                   REGION "INCREMENT FIRST STATION"
                       #firstStn += "simKP8Count";
                   END_REGION

                   REGION "UPPER LIMIT ROLL OVER"
                       IF #firstStn > "STATION_COUNT" THEN
                           #firstStn -= "STATION_COUNT" + 1;
                       END_IF;
                   END_REGION

               END_IF;
           END_REGION

           REGION "NEXT GROUP CHANGE DETECTION"
               #old.nextGrp := #currentBtn;
           END_REGION

       END_REGION

       REGION "PROCESS PREVIOUS GROUP PRESS"

           REGION "COPY TO LOCAL"
               #currentBtn := #simStations.up.actuate;
               #oldBtn := #old.prevGrp;
           END_REGION

           REGION "FALLING EDGE OF PREVIOUS GROUP"
               IF NOT #currentBtn AND #oldBtn THEN

                   REGION "DECREMENT FIRST STATION"
                       #firstStn -= "simKP8Count";
                   END_REGION

                   REGION "LOWER LIMIT ROLL OVER"
                       IF #firstStn < 0 THEN
                           #firstStn += "STATION_COUNT" + 1;
                       END_IF;
                   END_REGION

               END_IF;
           END_REGION

           REGION "PREVIOUS GROUP CHANGE DETECTION"
               #old.prevGrp := #currentBtn;
           END_REGION

       END_REGION

   END_REGION

   REGION "FOR EACH BUTTON"
       FOR #i := 0 TO 11 DO

           REGION "CALCULATE POINTER"
               #pStn := #i + #firstStn;
               #pSim := #i;
           END_REGION

           REGION "UPPER LIMIT ROLL OVER"
               IF #pStn > "STATION_COUNT" THEN
                   #pStn := #firstStn + #i - "STATION_COUNT" - 1;
               END_IF;
           END_REGION

           REGION "COPY TO LOCAL"
               #kp8Color := #stns.stn[#pStn].wipCmpts.ioData.kp8.tempOut;
           END_REGION

           REGION "LABEL STATIONS"

               REGION "DETERMINE LINE LABEL"
                   #label := #stns.stn[#pStn].id.lineName;
                   IF #label = #volvo16 THEN
                       #label := WSTRING#'V16';
                   END_IF;
               END_REGION

               REGION "DETERMINE DROP ZONE LABEL"
                   #intBox := USINT_TO_INT(#stns.stn[#pStn].id.dropZone);
                   IF #intBox <= 9 THEN
                       #dzLabel := CONCAT_WSTRING(IN1 := #lead0,
                                                  IN2 := "Strip Sign"(INT_TO_WSTRING(#intBox)));
                   END_IF;
                   IF #intBox >= 10 THEN
                       #dzLabel := "Strip Sign"(INT_TO_WSTRING(#intBox));
                   END_IF;
               END_REGION

               REGION "WRITE LABEL"
                   #label := CONCAT_WSTRING(IN1 := #label,
                                            IN2 := #space,
                                            IN3 := #dzLabel);
                   #simStations.me[#pSim].stn.label := #label;
               END_REGION

           END_REGION

           REGION "ANIMATE STATION LABEL"
               #simStations.me[#pSim].stn.animate := "GRAY_BACKGROUND";
           END_REGION

           REGION "FOR EACH BUTTON"
               FOR #j := 0 TO "STATION_BUTTON_COUNT" DO

                   REGION "COLOR BUTTONS"
                       #animate := "KP8 Driver: HMI Emulator: Animation"(kp8Color := #kp8Color,
                                                                btnNumber := #j);
                       #simStations.me[#pSim].btn.animate[#j] := #animate;
                   END_REGION

                   REGION "WRITE BUTTON LABELS"
                       #intBox := "Pointer Calc: KP8 Labels"(#j);
                       #label := "Strip Sign"(INT_TO_WSTRING(#intBox));
                       #simStations.me[#pSim].btn.labels[#j] := #label;
                   END_REGION

               END_FOR;
           END_REGION

       END_FOR;
   END_REGION

   REGION "SAVE FIRST STATION"
       #simStations.firstStn := #firstStn;
   END_REGION

   REGION "ANIMATE NEXT GROUP PRESS"
       #simStations.down.animate := "Bool.Animate"(true_color := "GREEN_LIGHT_BACKGROUND",
                                                   false_color := "GRAY_BACKGROUND",
                                                   evaluation_signal := #simStations.down.actuate);
   END_REGION

   REGION "ANIMATE PREV GROUP PARESS"
       #simStations.up.animate := "Bool.Animate"(true_color := "GREEN_LIGHT_BACKGROUND",
                                                 false_color := "GRAY_BACKGROUND",
                                                 evaluation_signal := #simStations.up.actuate);
   END_REGION
END_FUNCTION_BLOCK

FUNCTION "Sim: to Global" : Void   // FC23, SCL
{ S7_Optimized_Access := 'TRUE' }
VERSION : 0.1
   VAR_INPUT
      simStns : "Simulated Stations";
   END_VAR
   VAR_IN_OUT
      stations : "Station: All Stations";
   END_VAR
   VAR_TEMP
      i : Int;
      j : Int;
      pSim : Int;
      pStn : Int;
   END_VAR
BEGIN
   REGION "COPY TO LOCAL"
       // #btnCount := "btnCount";
       // #firstStn := #simStns.firstStn;
       // #simKP8Count := "simKP8Count";
       // #stnCount := "stnCount";
   END_REGION

   REGION "FOR EACH STATION"
       FOR #i := 0 TO "simKP8Count" DO

           REGION "CALCULATE POINTER"
               #pStn := #i + #simStns.firstStn;
               #pSim := #i;
           END_REGION

           REGION "UPPER LIMIT ROLL OVER"
               IF #pStn > "STATION_COUNT" THEN
                   #pStn := #simStns.firstStn + #i - "STATION_COUNT" - 1;
               END_IF;
           END_REGION

           REGION "COPY SIMULATED PRESSES"
               #stations.stn[#pStn].wipCmpts.ioData.kp8.input.%B1 := #simStns.me[#pSim].btn.actuate;
           END_REGION

       END_FOR;
   END_REGION
END_FUNCTION

FUNCTION "Sim: KP8 Animations" : Word   // FC84, SCL
{ S7_Optimized_Access := 'TRUE' }
VERSION : 0.1
   VAR_INPUT
      pbs : DWord;
   END_VAR
   VAR_TEMP
      ret : Word;
   END_VAR
BEGIN
   #"Sim: KP8 Animations".%B1 := #pbs.%B0;
   #"Sim: KP8 Animations".%B0 := #pbs.%B1;
END_FUNCTION

// folder: Linked List

FUNCTION_BLOCK "Linked List"   // FB29, SCL
{ S7_Optimized_Access := 'TRUE' }
VERSION : 0.1
   VAR_IN_OUT
      interface : "Linked List: Method Interface";
   END_VAR
   VAR
      list : "Linked List: List";
   END_VAR
   VAR CONSTANT
      TERMINAL_BEHAVIOR : String := 'open';
   END_VAR
BEGIN
   REGION "APPEND"
       IF #interface.append.in.request THEN
           "Linked List: Append"(terminal_behavior := #TERMINAL_BEHAVIOR,
                                 commands := #interface.append,
                                 list := #list);
       END_IF;
   END_REGION

   REGION "DELETE"
       IF #interface.delete.in.request THEN
           "Linked List: Delete"(commands := #interface.delete,
                                 list := #list);
       END_IF;
   END_REGION

   REGION "DISPLAY"
       IF #interface.display.in.request THEN
           "Linked List: Display"(commands := #interface.display,
                                  list := #list);
       END_IF;
   END_REGION

   REGION "INSERT"
       IF #interface.insert.in.request THEN
           "Linked List: Insert"(terminal_behavior := #TERMINAL_BEHAVIOR,
                                 commands := #interface.insert,
                                 list := #list);
       END_IF;
   END_REGION

   REGION "RESET"
       IF #interface.reset.in.request THEN
           "Linked List: Reset"(commands := #interface.reset,
                                list := #list);
       END_IF;
   END_REGION

   REGION "REVERSE"
       IF #interface.reverse.in.request THEN
           "Linked List: Reverse"(commands := #interface.reverse,
                                  list := #list);
       END_IF;
   END_REGION

   REGION "SEARCH"
       IF #interface.search.in.request THEN
           "Linked List: Search"(commands := #interface.search,
                                 list := #list);
       END_IF;
   END_REGION
END_FUNCTION_BLOCK

FUNCTION "Linked List: Private: Clear Node" : Void   // FC156, SCL
{ S7_Optimized_Access := 'TRUE' }
VERSION : 0.1
   VAR_IN_OUT
      node : "Linked List: Node";
   END_VAR
   VAR_TEMP
      ret : "Linked List: Node";
   END_VAR
BEGIN
   #ret.meta.key := "NULL_TOKEN";
   #ret.meta.next := "NULL_TOKEN";
   #node := #ret;
END_FUNCTION

FUNCTION "Linked List: Private: Get Head" : "Linked List: Node"   // FC157, SCL
{ S7_Optimized_Access := 'TRUE' }
VERSION : 0.1
   VAR_INPUT
      list : "Linked List: List";
   END_VAR
   VAR_TEMP
      pointer_list : DInt;
      ret : "Linked List: Node";
   END_VAR
BEGIN
   FOR #pointer_list := 0 TO "LINKED_LIST_LENGTH" DO
       IF #list.me[#pointer_list].meta.is_head THEN
           #ret := #list.me[#pointer_list];
           EXIT;
       END_IF;
   END_FOR;
   #"Linked List: Private: Get Head" := #ret;
END_FUNCTION

FUNCTION "Linked List: Private: Before" : Void   // FC158, SCL
{ S7_Optimized_Access := 'TRUE' }
VERSION : 0.1
   VAR_IN_OUT
      next_node : "Linked List: Node";   // next_node goes after node
      node : "Linked List: Node";   // node goes before next_node
   END_VAR
BEGIN
   #node.meta.next := #next_node.meta.key;
   IF #next_node.meta.is_head THEN
       #next_node.meta.is_head := FALSE;
       #node.meta.is_head := TRUE;
   END_IF;
END_FUNCTION

FUNCTION "Linked List: Private: Tail Swap" : Void   // FC159, SCL
{ S7_Optimized_Access := 'TRUE' }
VERSION : 0.1
   VAR_IN_OUT
      new_tail : "Linked List: Node";
      old_tail : "Linked List: Node";
   END_VAR
BEGIN
   #new_tail.meta.is_tail := TRUE;
   #old_tail.meta.is_tail := FALSE;
END_FUNCTION

FUNCTION "Linked List: Private: Head Swap" : Void   // FC160, SCL
{ S7_Optimized_Access := 'TRUE' }
VERSION : 0.1
   VAR_IN_OUT
      new_head : "Linked List: Node";
      old_head : "Linked List: Node";
   END_VAR
BEGIN
   #new_head.meta.is_head := TRUE;
   #old_head.meta.is_head := FALSE;
END_FUNCTION

FUNCTION "Linked List: Private: Get Next" : "Linked List: Node"   // FC161, SCL
{ S7_Optimized_Access := 'TRUE' }
VERSION : 0.1
   VAR_INPUT
      current : "Linked List: Node";
      list : "Linked List: List";
   END_VAR
   VAR_TEMP
      ret : "Linked List: Node";
   END_VAR
BEGIN
   "Linked List: Private: Clear Node"(#ret);
   IF #list.me[#current.meta.key].meta.next <> "NULL_TOKEN" THEN
       #ret := #list.me[#current.meta.next];
   END_IF;
   #"Linked List: Private: Get Next" := #ret;
END_FUNCTION

FUNCTION "Linked List: Private: Get Previous" : "Linked List: Node"   // FC162, SCL
{ S7_Optimized_Access := 'TRUE' }
VERSION : 0.1
   VAR_INPUT
      current : "Linked List: Node";
      list : "Linked List: List";
   END_VAR
   VAR_TEMP
      list_pointer : DInt;
      ret : "Linked List: Node";
   END_VAR
BEGIN
   "Linked List: Private: Clear Node"(#ret);
   FOR #list_pointer := 0 TO "LINKED_LIST_LENGTH" DO
       IF #list.me[#list_pointer].meta.next = #current.meta.key THEN
           #ret := #list.me[#list_pointer];
           EXIT;
       END_IF;
   END_FOR;
   #"Linked List: Private: Get Previous" := #ret;
END_FUNCTION

FUNCTION "Linked List: Private: After" : Void   // FC163, SCL
{ S7_Optimized_Access := 'TRUE' }
VERSION : 0.1
   VAR_IN_OUT
      node : "Linked List: Node";
      previous_node : "Linked List: Node";
   END_VAR
BEGIN
   #node.meta.next := #previous_node.meta.next;
   #previous_node.meta.next := #node.meta.key;
   IF #previous_node.meta.is_tail THEN
       #previous_node.meta.is_tail := FALSE;
       #node.meta.is_tail := TRUE;
   END_IF;
END_FUNCTION

FUNCTION "Linked List: Private: Head an Empty List" : Void   // FC164, SCL
{ S7_Optimized_Access := 'TRUE' }
VERSION : 0.1
   VAR_INPUT
      data : "Linked List: Node: Data";
      terminal_behavior : String;   // 'open': head's previous and tail's next are null nodes; 'closed': head's previous is tail, tail's next is head
   END_VAR
   VAR_IN_OUT
      list : "Linked List: List";
   END_VAR
BEGIN
   #list.me[0].data := #data;
   #list.me[0].meta.key := 0;
   IF #terminal_behavior = 'open' THEN
       #list.me[0].meta.next := "NULL_TOKEN";
   END_IF;
   IF #terminal_behavior = 'closed' THEN
       #list.me[0].meta.next := 0;
   END_IF;
   #list.me[0].meta.is_head := TRUE;
   #list.me[0].meta.is_tail := TRUE;
END_FUNCTION

FUNCTION "Linked List: Private: Is Empty" : Bool   // FC165, SCL
{ S7_Optimized_Access := 'TRUE' }
VERSION : 0.1
   VAR_INPUT
      list : "Linked List: List";
   END_VAR
   VAR_TEMP
      pointer_list : DInt;
      ret : Bool;
   END_VAR
BEGIN
   #ret := TRUE;
   FOR #pointer_list := 0 TO "LINKED_LIST_LENGTH" DO
       IF #list.me[#pointer_list].meta.key <> "NULL_TOKEN" THEN
           #ret := FALSE;
           EXIT;
       END_IF;
   END_FOR;
   #"Linked List: Private: Is Empty" := #ret;
END_FUNCTION

FUNCTION "Linked List: Private: Get Tail" : "Linked List: Node"   // FC166, SCL
{ S7_Optimized_Access := 'TRUE' }
VERSION : 0.1
   VAR_IN_OUT
      list : "Linked List: List";
   END_VAR
   VAR_TEMP
      pointer_list : Int;
      next_node : UInt;
      ret : "Linked List: Node";
   END_VAR
BEGIN
   FOR #pointer_list := 0 TO "LINKED_LIST_LENGTH" DO
       IF #list.me[#pointer_list].meta.is_tail THEN
           #ret := #list.me[#pointer_list];
           EXIT;
       END_IF;
   END_FOR;
   #"Linked List: Private: Get Tail" := #ret;
END_FUNCTION

FUNCTION "Linked List: Private: Is Full" : Bool   // FC167, SCL
{ S7_Optimized_Access := 'TRUE' }
VERSION : 0.1
   VAR_INPUT
      list : "Linked List: List";
   END_VAR
   VAR_TEMP
      pointer_list : DInt;
      ret : Bool;
   END_VAR
BEGIN
   #ret := TRUE;
   FOR #pointer_list := 0 TO "LINKED_LIST_LENGTH" DO
       IF #list.me[#pointer_list].meta.key = "NULL_TOKEN" THEN
           #ret := FALSE;
           EXIT;
       END_IF;
   END_FOR;
   #"Linked List: Private: Is Full" := #ret;
END_FUNCTION

FUNCTION "Linked List: Private: Next Empty Node" : DInt   // FC168, SCL
{ S7_Optimized_Access := 'TRUE' }
VERSION : 0.1
   VAR_IN_OUT
      list : "Linked List: List";
   END_VAR
   VAR_TEMP
      node : "Linked List: Node";
      pointer_list : Int;
      ret : DInt;
   END_VAR
BEGIN
   #ret := "NULL_TOKEN";
   FOR #pointer_list := 0 TO "LINKED_LIST_LENGTH" DO
       IF #list.me[#pointer_list].meta.key = "NULL_TOKEN" THEN
           #ret := INT_TO_DINT(#pointer_list);
           EXIT;
       END_IF;
   END_FOR;
   #"Linked List: Private: Next Empty Node" := #ret;
END_FUNCTION

FUNCTION "Linked List: Append" : Void   // FC169, SCL
{ S7_Optimized_Access := 'TRUE' }
VERSION : 0.1
   VAR_INPUT
      terminal_behavior : String;
   END_VAR
   VAR_IN_OUT
      commands : "Linked List: Method Interface: Append";
      list : "Linked List: List";
   END_VAR
   VAR_TEMP
      clear_commands : "Linked List: Method Interface: Append";
      head : "Linked List: Node";
      pointer_new_node : DInt;
      tail : "Linked List: Node";
   END_VAR
   VAR CONSTANT
      no_error : String := 'no error';
      list_full : String := 'appended to full list';
      no_tail_found : String := 'no tail found while trying to append';
      appended_as_head : String := 'appended as head of list';
   END_VAR
BEGIN
   REGION "NOTES"
       (*
       Append adds a node to the end of the list.
       Last edit: 2021-10-05
       *)
   END_REGION

   REGION "APPEND TO FULL LIST"
       IF "Linked List: Private: Is Full"(#list) THEN
           #commands := #clear_commands;
           #commands.out.error := TRUE;
           #commands.out.error_message := #list_full;
           RETURN;
       END_IF;
   END_REGION

   REGION "APPEND TO EMPTY LIST"
       IF "Linked List: Private: Is Empty"(#list) THEN
           "Linked List: Private: Head an Empty List"(data := #commands.in.data,
                                                      terminal_behavior := #terminal_behavior,
                                                      list := #list);
           #commands := #clear_commands;
           #commands.out.done := TRUE;
           #commands.out.error_message := #appended_as_head;
           RETURN;
       END_IF;
   END_REGION

   REGION "FIND TAIL"
       #tail := "Linked List: Private: Get Tail"(#list);
   END_REGION

   REGION "EXIT CONDITION: TAIL NOT FOUND"
       IF #tail.meta.key = "NULL_TOKEN" THEN
           #commands := #clear_commands;
           #commands.out.error := TRUE;
           #commands.out.error_message := #no_tail_found;
           RETURN;
       END_IF;
   END_REGION

   REGION "FIND FIRST NULL"
       #pointer_new_node := "Linked List: Private: Next Empty Node"(#list);
   END_REGION

   REGION "APPENDED NODE IS AFTER TAIL"
       #list.me[#pointer_new_node].data := #commands.in.data;
       #list.me[#pointer_new_node].meta.key := #pointer_new_node;
       "Linked List: Private: After"(node := #list.me[#pointer_new_node],
                                     previous_node := #list.me[#tail.meta.key]);
   END_REGION

   REGION "EXIT CONDITION: SUCCESS"
       #commands := #clear_commands;
       #commands.out.done := TRUE;
       #commands.out.error_message := #no_error;
   END_REGION
END_FUNCTION

FUNCTION "Linked List: Delete" : Void   // FC170, SCL
{ S7_Optimized_Access := 'TRUE' }
VERSION : 0.1
   VAR_IN_OUT
      commands : "Linked List: Method Interface: Delete";
      list : "Linked List: List";
   END_VAR
   VAR_TEMP
      blank_node : "Linked List: Node";
      clear_commands : "Linked List: Method Interface: Delete";
      current : "Linked List: Node";
      found : Bool;
      next : "Linked List: Node";
      pointer_list : DInt;
      previous : "Linked List: Node";
      search_commands : "Linked List: Method Interface: Search";
   END_VAR
   VAR CONSTANT
      no_error : String := 'no error';
      delete_from_empty : String := 'deleted from an empty list.';
   END_VAR
BEGIN
   REGION "EXIT CONDITION: LIST IS EMPTY"
       IF "Linked List: Private: Is Empty"(#list) THEN
           #commands := #clear_commands;
           #commands.out.error := TRUE;
           #commands.out.error_message := #delete_from_empty;
       END_IF;
   END_REGION

   REGION "DELETE"
       #current := #commands.in.node;
       #previous := "Linked List: Private: Get Previous"(current := #current,
                                                         list := #list);
       #next := "Linked List: Private: Get Next"(current := #current,
                                                 list := #list);
       IF #current.meta.is_head AND NOT #current.meta.is_tail THEN
           "Linked List: Private: Head Swap"(new_head := #list.me[#next.meta.key],
                                             old_head := #list.me[#current.meta.key]);
       END_IF;
       IF NOT #current.meta.is_head AND #current.meta.is_tail THEN
           "Linked List: Private: Tail Swap"(new_tail := #list.me[#previous.meta.key],
                                             old_tail := #list.me[#current.meta.key]);
       END_IF;
       IF NOT #current.meta.is_head THEN
           #list.me[#previous.meta.key].meta.next := #next.meta.key;
       END_IF;
       "Linked List: Private: Clear Node"(#list.me[#current.meta.key]);
   END_REGION

   REGION "COMMANDS OUT"
       #commands := #clear_commands;
       #commands.out.done := TRUE;
       #commands.out.error_message := #no_error;
   END_REGION
END_FUNCTION

FUNCTION "Linked List: Search" : Void   // FC171, SCL
{ S7_Optimized_Access := 'TRUE' }
VERSION : 0.1
   VAR_IN_OUT
      commands : "Linked List: Method Interface: Search";
      list : "Linked List: List";
   END_VAR
   VAR_TEMP
      clear_commands : "Linked List: Method Interface: Search";
      found : Bool;
      pointer_list : DInt;
   END_VAR
   VAR CONSTANT
      no_error : String := 'no error';
      searched_empty_list : String := 'searched empty list';
   END_VAR
BEGIN
   REGION "EXIT CONDITION: SEARCHED EMPTY LIST"
       IF "Linked List: Private: Is Empty"(#list) THEN
           #commands := #clear_commands;
           #commands.out.not_found := TRUE;
           #commands.out.error := TRUE;
           #commands.out.error_message := #searched_empty_list;
           RETURN;
       END_IF;
   END_REGION

   REGION "SEARCH"
       FOR #pointer_list := 0 TO "LINKED_LIST_LENGTH" DO
           IF #list.me[#pointer_list].data = #commands.in.data THEN
               #found := TRUE;
               EXIT;
           END_IF;
       END_FOR;
   END_REGION

   REGION "FOUND"
       IF #found THEN
           #commands := #clear_commands;
           #commands.out.done := TRUE;
           #commands.out.found := TRUE;
           #commands.out.returned_node := #list.me[#pointer_list];
           #commands.out.error_message := #no_error;
           RETURN;
       END_IF;
   END_REGION

   REGION "NOT FOUND"
       IF NOT #found THEN
           #commands := #clear_commands;
           #commands.out.done := TRUE;
           #commands.out.not_found := TRUE;
           RETURN;
       END_IF;
   END_REGION
END_FUNCTION

FUNCTION "Linked List: Display" : Void   // FC172, SCL
{ S7_Optimized_Access := 'TRUE' }
VERSION : 0.1
   VAR_IN_OUT
      commands : "Linked List: Method Interface: Display";
      list : "Linked List: List";
   END_VAR
   VAR_TEMP
      clear_commands : "Linked List: Method Interface: Display";
   END_VAR
BEGIN
   #commands := #clear_commands;
   #commands.out.list := #list;
   #commands.out.done := TRUE;
END_FUNCTION

FUNCTION "Linked List: Insert" : Void   // FC173, SCL
{ S7_Optimized_Access := 'TRUE' }
VERSION : 0.1
   VAR_INPUT
      terminal_behavior : String;
   END_VAR
   VAR_IN_OUT
      commands : "Linked List: Method Interface: Insert";
      list : "Linked List: List";
   END_VAR
   VAR_TEMP
      clear_commands : "Linked List: Method Interface: Insert";
      current : "Linked List: Node";
      next_empty_node_index : DInt;
      previous : "Linked List: Node";
      next : "Linked List: Node";
   END_VAR
   VAR CONSTANT
      no_error : String := 'no error';
      inserted_into_full : String := 'attempted to insert into full list. delete a node and try again.';
      appended_as_head : String := 'appended as head of list';
   END_VAR
BEGIN
   REGION "EXIT CONDITION: INSERTED INTO FULL LIST"
       IF "Linked List: Private: Is Full"(#list) THEN
           #commands := #clear_commands;
           #commands.out.error := TRUE;
           #commands.out.error_message := #inserted_into_full;
           RETURN;
       END_IF;
   END_REGION

   REGION "EXIT CONDITION: INSERTED INTO EMPTY LIST"
       IF "Linked List: Private: Is Empty"(#list) THEN
           "Linked List: Private: Head an Empty List"(data := #commands.in.data,
                                                      terminal_behavior := #terminal_behavior,
                                                      list := #list);
           #commands := #clear_commands;
           #commands.out.error := TRUE;
           #commands.out.error_message := #appended_as_head;
           RETURN;
       END_IF;
   END_REGION

   REGION "GET INDEX OF NEXT EMPTY NODE"
       #next_empty_node_index := "Linked List: Private: Next Empty Node"(#list);
   END_REGION

   REGION "PREVIOUS, CURRENT, AND NEXT NODES"
       #current := #commands.in.target_node;
       #previous := "Linked List: Private: Get Previous"(current := #current,
                                                         list := #list);
       #next := #current;
   END_REGION

   REGION "INSERT BEFORE TARGET NODE"
       // new node's data becomes command data
       #list.me[#next_empty_node_index].data := #commands.in.data;
       // new node's key becomes array index
       #list.me[#next_empty_node_index].meta.key := #next_empty_node_index;
       // shorten name for indexing
       #current := #list.me[#next_empty_node_index];
       // insert
       IF NOT #next.meta.is_head THEN
           "Linked List: Private: After"(node := #list.me[#current.meta.key],
                                         previous_node := #list.me[#previous.meta.key]);
       END_IF;
       "Linked List: Private: Before"(next_node := #list.me[#next.meta.key],
                                      node := #list.me[#current.meta.key]);
   END_REGION

   REGION "COMMANDS OUT"
       #commands := #clear_commands;
       #commands.out.done := TRUE;
       #commands.out.error_message := #no_error;
   END_REGION
END_FUNCTION

FUNCTION "Linked List: Reverse" : Void   // FC174, SCL
{ S7_Optimized_Access := 'TRUE' }
VERSION : 0.1
   VAR_IN_OUT
      commands : "Linked List: Method Interface: Reverse";
      list : "Linked List: List";
   END_VAR
   VAR_TEMP
      clear_commands : "Linked List: Method Interface: Reverse";
      current : "Linked List: Node";
      next : "Linked List: Node";
      previous : "Linked List: Node";
      null_node : "Linked List: Node";
   END_VAR
   VAR CONSTANT
      no_error : String := 'no error';
      reversed_empty_list : String := 'reversed empty list';
   END_VAR
BEGIN
   IF "Linked List: Private: Is Empty"(#list) THEN
       #commands := #clear_commands;
       #commands.out.error := TRUE;
       #commands.out.error_message := #reversed_empty_list;
       RETURN;
   END_IF;

   "Linked List: Private: Clear Node"(#null_node);
   #previous := #null_node;
   #current := "Linked List: Private: Get Head"(#list);
   #list.me[#current.meta.key].meta.is_head := FALSE;
   #list.me[#current.meta.key].meta.is_tail := TRUE;
   WHILE #current.meta.next <> "NULL_TOKEN" DO
       #next := #list.me[#current.meta.next];
       #list.me[#current.meta.key].meta.next := #previous.meta.key;
       #previous := #current;
       #current := #next;
       #list.me[#current.meta.key].meta.is_head := FALSE;
       #list.me[#current.meta.key].meta.is_tail := FALSE;
   END_WHILE;
   #list.me[#current.meta.key].meta.next := #previous.meta.key;
   #list.me[#current.meta.key].meta.is_head := TRUE;
   #list.me[#current.meta.key].meta.is_tail := FALSE;

   #commands := #clear_commands;
   #commands.out.done := TRUE;
   #commands.out.error_message := #no_error;
END_FUNCTION

FUNCTION "Linked List: Reset" : Void   // FC175, SCL
{ S7_Optimized_Access := 'TRUE' }
VERSION : 0.1
   VAR_IN_OUT
      commands : "Linked List: Method Interface: Reset";
      list : "Linked List: List";
   END_VAR
   VAR_TEMP
      blank_node : "Linked List: Node";
      list_pointer : DInt;
      clear_commands : "Linked List: Method Interface: Reset";
   END_VAR
BEGIN
   FOR #list_pointer := 0 TO "LINKED_LIST_LENGTH" DO
       "Linked List: Private: Clear Node"(#list.me[#list_pointer]);
   END_FOR;
   #commands := #clear_commands;
   #commands.out.done := TRUE;
END_FUNCTION

// folder: OBs

ORGANIZATION_BLOCK "Rack or station failure"   // OB86, LAD, RackStationFailure
{ S7_Optimized_Access := 'TRUE' }
VERSION : 0.1
   VAR_INPUT
      LADDR : Hw_Device;   // Hardware identifier
      Event_Class : Byte;   // Event class
      Fault_ID : Byte;   // Fault identifier
   END_VAR
BEGIN
END_ORGANIZATION_BLOCK

ORGANIZATION_BLOCK "Startup"   // OB100, LAD, Startup
TITLE = "Complete Restart"
{ S7_Optimized_Access := 'TRUE' }
VERSION : 0.1
   VAR_INPUT
      LostRetentive : Bool;   // True if retentive data are lost
      LostRTC : Bool;   // True if date and time are lost
   END_VAR
BEGIN

REGION Network 1 (SCL): HMI STATION INITIALIZATION
END_REGION
END_ORGANIZATION_BLOCK

ORGANIZATION_BLOCK "Programming error"   // OB121, LAD, ProgrammingError
{ S7_Optimized_Access := 'TRUE' }
VERSION : 0.1
   VAR_INPUT
      BlockNr : UInt;   // Number of causing block
      Reaction : USInt;   // 0:ignore, 1:substitute, 2:skip
      Fault_ID : Byte;   // Fault identifier
      BlockType : USInt;   // 16#01:OB, 16#02:FC, 16#03:FB, 16#04:SFC, 16#05:SFB, 16#06:DB: Type of block causing the error
      Area : USInt;   // Area where the error occured
      DBNr : DB_ANY;   // DB number if Area = DB or DI
      Csg_OBNr : OB_Any;   // Number of OB causing the error
      Csg_Prio : USInt;   // Priority of OB causing the error
      Width : USInt;   // 0:bit, 1:byte, 2:word, 3:dword, 4:lword
   END_VAR
BEGIN
END_ORGANIZATION_BLOCK

ORGANIZATION_BLOCK "IO access error"   // OB122, LAD, IOAccessError
{ S7_Optimized_Access := 'TRUE' }
VERSION : 0.1
   VAR_INPUT
      BlockNr : UInt;   // Number of causing block
      Reaction : USInt;   // 0:ignore, 1:substitute, 2:skip
      Fault_ID : Byte;   // 16#42:reading, 16#43:writing
      BlockType : USInt;   // 16#01:OB, 16#02:FC, 16#03:FB, 16#04:SFC, 16#05:SFB, 16#06:DB: Type of block causing the error
      Area : USInt;   // 16#81:I, 16#82:Q: IO area where the IOaccess error occured
      DBNr : DB_ANY;   // Reserved for system
      Csg_OBNr : OB_Any;   // Number of OB causing the error
      Csg_Prio : USInt;   // Priority of OB causing the error
      Width : USInt;   // 0:bit, 1:byte, 2:word, 3:dword, 4:lword
   END_VAR
BEGIN
END_ORGANIZATION_BLOCK

// folder: Order/States

FUNCTION_BLOCK "Order State"   // FB2, SCL
{ S7_Optimized_Access := 'TRUE' }
VERSION : 0.1
   VAR_INPUT
      pnLib : "Recipe: PN Text Library";
   END_VAR
   VAR_IN_OUT
      stns : "Station: All Stations";
   END_VAR
   VAR_TEMP
      pStn : Int;
      pBtn : Int;
      stn : "Station: Single Station";
   END_VAR
BEGIN
   REGION "FOR EACH STATION"
       FOR #pStn := 0 TO "STATION_COUNT" DO

           REGION "FOR EACH BUTTON"
               FOR #pBtn := 0 TO "STATION_BUTTON_COUNT" DO

                   REGION "POPULATE CURRENT STATION"
                       #stn := #stns.stn[#pStn];
                   END_REGION

                   REGION "INITIALIZE STATE"
                       "Order State: Initialize State"(newParams := #stn.wipCmpts.flags.newPN,
                                                       pnGood := #stn.wipCmpts.flags.pnGood[#pBtn],
                                                       state := #stn.wipCmpts.orderState[#pBtn]);
                   END_REGION

                   REGION "ENTER IDLE"
                       "Order State: Enter Idle"(btnFalling := #stn.wipCmpts.kp8Logical.falling.btn[#pBtn],
                                                 state := #stn.wipCmpts.orderState[#pBtn]);
                   END_REGION

                   REGION "ENTER REQUESTED"
                       "Order State: Enter Requested"(btnRising := #stn.wipCmpts.kp8Logical.rising.btn[#pBtn],
                                                      state := #stn.wipCmpts.orderState[#pBtn]);
                   END_REGION

                   REGION "ENTER REQUESTED CRITICAL"
                       "Order State: Enter Requested Critical"(timerVal := #stn.wipCmpts.timers.remaining[#pBtn],
                                                               state := #stn.wipCmpts.orderState[#pBtn]);
                   END_REGION

                   REGION "ENTER REQUESTED EXPIRED"
                       "Order State: Enter Requested Expired"(timerVal := #stn.wipCmpts.timers.remaining[#pBtn],
                                                              state := #stn.wipCmpts.orderState[#pBtn]);
                   END_REGION

                   REGION "SAVE CURRENT STATION"
                       #stns.stn[#pStn] := #stn;
                   END_REGION

               END_FOR;
           END_REGION

       END_FOR;
   END_REGION
END_FUNCTION_BLOCK

FUNCTION "Order State: Enter Idle" : Void   // FC6, SCL
{ S7_Optimized_Access := 'TRUE' }
VERSION : 0.1
   VAR_INPUT
      btnFalling : Bool;
   END_VAR
   VAR_IN_OUT
      state : Int;
   END_VAR
BEGIN
   IF #btnFalling THEN
       #state := "idle";
   END_IF;
END_FUNCTION

FUNCTION "Order State: Enter Requested" : Void   // FC7, SCL
{ S7_Optimized_Access := 'TRUE' }
VERSION : 0.1
   VAR_INPUT
      btnRising : Bool;
   END_VAR
   VAR_IN_OUT
      state : Int;
   END_VAR
BEGIN
   IF #state = "idle" THEN
       IF #btnRising THEN
           #state := "requested";
       END_IF;
   END_IF;
END_FUNCTION

FUNCTION "Order State: Initialize State" : Void   // FC10, SCL
{ S7_Optimized_Access := 'TRUE' }
VERSION : 0.1
   VAR_INPUT
      newParams : Bool;
      pnGood : Bool;
   END_VAR
   VAR_IN_OUT
      state : Int;
   END_VAR
BEGIN
   REGION "ON NEW PARAMETERS"
       IF #newParams THEN

           REGION "ON VALID PN" 
               IF #pnGood THEN

                   REGION "INITIALIZE STATE"
                       #state := BOOL_TO_INT(#pnGood);
                   END_REGION

               END_IF;
           END_REGION

       END_IF;
   END_REGION
END_FUNCTION

FUNCTION "Order State: Enter Requested Critical" : Void   // FC16, SCL
{ S7_Optimized_Access := 'TRUE' }
VERSION : 0.1
   VAR_INPUT
      timerVal : Real;
   END_VAR
   VAR_IN_OUT
      state : Int;
   END_VAR
   VAR_TEMP
      temp : Real;
   END_VAR
BEGIN
   IF #state = "requested" THEN
       IF #timerVal > 0.0 AND #timerVal <= "tCritical" THEN
           #state := "requestedCrit";
       END_IF;
   END_IF;
END_FUNCTION

FUNCTION "Order State: Enter Requested Expired" : Void   // FC17, SCL
{ S7_Optimized_Access := 'TRUE' }
VERSION : 0.1
   VAR_INPUT
      timerVal : Real;
   END_VAR
   VAR_IN_OUT
      state : Int;
   END_VAR
BEGIN
   IF #state = "requestedCrit" THEN
       IF #timerVal <= -0.001 THEN
           #state := "requestedExp";
       END_IF;
   END_IF;
END_FUNCTION

// folder: Order/Timers

FUNCTION_BLOCK "Order Timer"   // FB6, SCL
{ S7_Optimized_Access := 'TRUE' }
VERSION : 0.1
   VAR_INPUT
      pnLib : "Recipe: PN Text Library";
   END_VAR
   VAR_IN_OUT
      stns : "Station: All Stations";
   END_VAR
   VAR
      rt : "Runtime Data";
   END_VAR
   VAR_TEMP
      pStn : Int;
      pBtn : Int;
   END_VAR
BEGIN
   REGION "RUNTIME CALL"
       #rt.elapsed := RUNTIME(#rt.mem);
       #rt.asReal := LREAL_TO_REAL(#rt.elapsed);
   END_REGION

   REGION "FOR EACH STATION"
       FOR #pStn := 0 TO "STATION_COUNT" DO

           REGION "FOR EACH BUTTON"
               FOR #pBtn := 0 TO "STATION_BUTTON_COUNT" DO

                   REGION "INITIALIZE TIMERS"
                       "Order Timer: Initialize"(pnLib := #pnLib,
                                                 pBtn := #pBtn,
                                                 stn := #stns.stn[#pStn]);
                   END_REGION

                   REGION "EXECUTE TIMERS"
                       "Order Timer: Timer Execution"(elapsedTime := #rt.asReal,
                                                      pBtn := #pBtn,
                                                      stn:=#stns.stn[#pStn],
                                                      timers := #stns.stn[#pStn].wipCmpts.timers);
                   END_REGION

               END_FOR;
           END_REGION

       END_FOR;
   END_REGION
END_FUNCTION_BLOCK

FUNCTION "Order Timer: Initialize" : Void   // FC8, SCL
{ S7_Optimized_Access := 'TRUE' }
VERSION : 0.1
   VAR_INPUT
      pnLib : "Recipe: PN Text Library";
      pBtn : Int;
   END_VAR
   VAR_IN_OUT
      stn : "Station: Single Station";
   END_VAR
   VAR_TEMP
      pnGood : Bool;
      default : Bool;
      clear : Bool;
   END_VAR
BEGIN
   REGION "ON PN CHANGE"
       IF #stn.wipCmpts.flags.newPN THEN

           REGION "INITIALIZE TO DEFAULT"

               REGION "EXECUTION VALIDATION"
                   #default := "Order Timer: Set to Default Check"(pnGood := #stn.wipCmpts.flags.pnGood[#pBtn],
                                                                   inSettingsScreen := #stn.wipCmpts.flags.inSettingsScreen,
                                                                   timerReset := #stn.wipCmpts.flags.resetTimer[#pBtn]);
               END_REGION

               REGION "ON VALIDATION"
                   IF #default THEN

                       REGION "SET DEFAULT TIME VALUE"
                           #stn.wipCmpts.timers.ptAllotted[#pBtn] := "tAllotted";
                           #stn.wipCmpts.timers.ptCritical[#pBtn] := "tCritical";
                       END_REGION

                   END_IF;
               END_REGION

           END_REGION

           REGION "INITIALIZE TO ZERO"

               REGION "EXECUTION VALIDATION"
                   #clear := "Order Timer: Set to Zero Check"(pnGood := #stn.wipCmpts.flags.pnGood[#pBtn],
                                                              inSettingsScreen := #stn.wipCmpts.flags.inSettingsScreen,
                                                              timerReset := #stn.wipCmpts.flags.resetTimer[#pBtn]);
               END_REGION

               REGION "ON VALIDATION"
                   IF #clear THEN

                       REGION "SET DEFAULT TIME VALUE"
                           #stn.wipCmpts.timers.ptAllotted[#pBtn] := 0.0;
                           #stn.wipCmpts.timers.ptCritical[#pBtn] := 0.0;
                       END_REGION

                   END_IF;
               END_REGION

           END_REGION

       END_IF;
   END_REGION
END_FUNCTION

FUNCTION "Order Timer: Timer Execution" : Void   // FC11, SCL
{ S7_Optimized_Access := 'TRUE' }
VERSION : 0.1
   VAR_INPUT
      elapsedTime : Real;
      pBtn : Int;
      stn : "Station: Single Station";
   END_VAR
   VAR_IN_OUT
      timers : "Station: Timers";
   END_VAR
BEGIN
   REGION "RUN CONDITIONS"
       CASE #stn.wipCmpts.orderState[#pBtn] OF

           "reset", "idle":
               IF #stn.flags.stateTransition[#pBtn] THEN
                   #timers.elapsed[#pBtn] := 0.0;
                   #timers.remaining[#pBtn] := 0.0;
               END_IF;

           "requested".."acknowledgedExp":
               #timers.elapsed[#pBtn] += #elapsedTime;
               #timers.remaining[#pBtn] := #timers.ptAllotted[#pBtn] - #timers.elapsed[#pBtn];

           ELSE:
               ;

       END_CASE;
   END_REGION
END_FUNCTION

FUNCTION "Order Timer: Set to Default Check" : Bool   // FC12, SCL
{ S7_Optimized_Access := 'TRUE' }
VERSION : 0.1
   VAR_INPUT
      pnGood : Bool;
      inSettingsScreen : Bool;
      timerReset : Bool;
   END_VAR
   VAR_TEMP
      ret : Bool;
   END_VAR
BEGIN
   REGION "ON VALID PN"
       #ret := #pnGood;
   END_REGION

   REGION "NOT WHILE IN SETTINGS SCREEN"
       IF #inSettingsScreen THEN
           #ret := FALSE;
       END_IF;
   END_REGION

   REGION "ON RESET REQUEST"
       #ret := #timerReset OR #ret;
   END_REGION

   REGION "RETURN"
       #"Order Timer: Set to Default Check" := #ret;
   END_REGION
END_FUNCTION

FUNCTION "Order Timer: Set to Zero Check" : Bool   // FC15, SCL
{ S7_Optimized_Access := 'TRUE' }
VERSION : 0.1
   VAR_INPUT
      pnGood : Bool;
      inSettingsScreen : Bool;
      timerReset : Bool;
   END_VAR
   VAR_TEMP
      ret : Bool;
   END_VAR
BEGIN
   REGION "ON VALID PN"
       #ret := NOT #pnGood;
   END_REGION

   REGION "NOT WHILE IN SETTINGS SCREEN"
       IF #inSettingsScreen THEN
           #ret := FALSE;
       END_IF;
   END_REGION

   REGION "ON RESET REQUEST"
       #ret := #timerReset OR #ret;
   END_REGION

   REGION "RETURN"
       #"Order Timer: Set to Zero Check" := #ret;
   END_REGION
END_FUNCTION

// folder: Part Request

FUNCTION_BLOCK "Part Request"   // FB7, SCL
{ S7_Optimized_Access := 'TRUE' }
VERSION : 0.1
   VAR_INPUT
      stns : "Station: All Stations";
      savedWips : "Recipe: HMI Stations Saved Wips";
      pnLib : "Recipe: PN Text Library";
   END_VAR
   VAR_IN_OUT
      dataTable : "Part Request Data";
   END_VAR
   VAR RETAIN
      pDataRow : Int;
   END_VAR
   VAR_TEMP
      address : DInt;
      addRequest : Bool;
      inTable : DInt;
      pStn : Int;
      pBtn : Int;
      pWip : Int;
      pRqstsRow : Int;
      removeRequest : Bool;
   END_VAR
BEGIN
   REGION "FOR EACH STATION"
       FOR #pStn := 0 TO "STATION_COUNT" DO

           REGION "FOR EACH BUTTON"
               FOR #pBtn := 0 TO "STATION_BUTTON_COUNT" DO

                   REGION "NEXT BUTTON ON NO TRANSITION"
                       IF NOT #stns.stn[#pStn].flags.stateTransition[#pBtn] THEN
                           GOTO NOSTNREQ;
                       END_IF;
                   END_REGION

                   REGION "GET ADDRESS"
                       #pWip := DINT_TO_INT(#stns.stn[#pStn].wipData.index);
                       #address := "Address.Set_Address"(pStn := #pStn, pBtn := #pBtn, pWip := #pWip);
                   END_REGION

                   REGION "CHECK FOR ENTRY IN DATA TABLE"
                       #inTable := "Part Request: Address in Table"(search := #address,
                                                                    dataTable := #dataTable);
                   END_REGION

                   REGION "ADD"

                       REGION "VALIDATE CONDITIONS"
                           #addRequest := "Part Request: Validate Add"(inTable := #inTable,
                                                                       orderState := #stns.stn[#pStn].wipCmpts.orderState[#pBtn]);
                       END_REGION

                       REGION "EXECUTE"
                           IF #addRequest THEN
                               #addRequest := FALSE;
                               #dataTable.row[#pDataRow] := #address;
                               "Row Pointer: Roll Over"(limit := "partReqDataRowCount",
                                                                "pointer" := #pDataRow);
                           END_IF;
                       END_REGION

                   END_REGION

                   REGION "REMOVE SINGLE STATION"

                       REGION "VALIDATE CONDITIONS: SINGLE"
                           #removeRequest := "Part Request: Validate Remove: Single"(inTable := #inTable,
                                                                                     orderState := #stns.stn[#pStn].wipCmpts.orderState[#pBtn]);
                       END_REGION

                       REGION "EXECUTE"
                           IF #removeRequest THEN
                               #removeRequest := FALSE;
                               #dataTable.row[#inTable] := -1;
                               "Part Request: Collapse Table"(#dataTable);
                               "Row Pointer: Post Collapse"(dataTable := #dataTable,
                                                            pDataRow := #pDataRow);
                           END_IF;
                       END_REGION

                   END_REGION

               NOSTNREQ:
                   ;
               END_FOR;
           END_REGION

       END_FOR;
   END_REGION


   (* REGION "REMOVE WIP STATIONS"                    
       FOR #pStn := 0 TO "hmiStnCount" DO
           FOR #pWip := 0 TO "wipCount" DO
               IF #savedWips.stn[#pStn].wip[#pWip].flags.clearWipRequest THEN
                   FOR #pBtn := 0 TO "btnCount" DO
                       #address := "Address: Set Address"(pBtn := #pBtn, pStn := #pStn, pWip := #pWip);
                       #inTable := "Part Request: Address in Table"(adrRequest := #address,
                                                                    dataTable := #dataTable);
                       #removeRequest := "Part Request: Validate Remove: WIP"(inTable := #inTable,
                                                                              clearWipRequest := #savedWips.stn[#pStn].wip[#pWip].flags.clearWipRequest);
                       IF #removeRequest THEN
                           #removeRequest := FALSE;
                           "Part Request: Remove"(pRow := #inTable,
                                                  dataTable := #dataTable);
                           "Part Request: Collapse Table"(#dataTable);
                           "Row Pointer: Post Collapse"(dataTable := #dataTable,
                                                        pDataRow := #pDataRow);
                       END_IF;
                   END_FOR;
               END_IF;
           END_FOR;
       END_FOR;
   END_REGION *)
END_FUNCTION_BLOCK

FUNCTION "Part Request: Address in Table" : DInt   // FC27, SCL
{ S7_Optimized_Access := 'TRUE' }
VERSION : 0.1
   VAR_INPUT
      search : DInt;
      dataTable : "Part Request Data";
   END_VAR
   VAR_TEMP
      ret : DInt;
      pRow : DInt;
   END_VAR
BEGIN
   REGION "DEFAULT RETURN"    
       #ret := -1;
   END_REGION

   REGION "CHECK TABLE"
       WHILE #dataTable.row[#pRow] <> #search AND #pRow <= "partReqDataRowCount" DO
           #pRow += 1;
       END_WHILE;
       IF #pRow <= "partReqDataRowCount" THEN
           #ret := #pRow;
       END_IF;
   END_REGION

   REGION "RETURN"
       #"Part Request: Address in Table" := #ret;
   END_REGION

   REGION "CALL READ VFD"
       ;
       ;
   END_REGION
END_FUNCTION

FUNCTION "Part Request: Validate Add" : Bool   // FC30, SCL
{ S7_Optimized_Access := 'TRUE' }
VERSION : 0.1
   VAR_INPUT
      inTable : DInt;
      orderState : Int;
   END_VAR
   VAR_TEMP
      ret : Bool;
   END_VAR
BEGIN
   IF #inTable = -1 THEN
       CASE #orderState OF
           "idle",
           "requestedCrit", "requestedExp",
           "ordered", "orderedCrit", "orderedExp",
           "acknowledged", "acknowledgedCrit", "acknowledgedExp":
               #ret := FALSE;
           "requested":
               #ret := TRUE;
       END_CASE;
   END_IF;
   #"Part Request: Validate Add" := #ret;
END_FUNCTION

FUNCTION "Part Request: Validate Remove: Single" : Bool   // FC41, SCL
{ S7_Optimized_Access := 'TRUE' }
VERSION : 0.1
   VAR_INPUT
      inTable : DInt;
      orderState : Int;
   END_VAR
   VAR_TEMP
      ret : Bool;
   END_VAR
BEGIN
   IF #inTable <> -1 THEN
       CASE #orderState OF
           "requested", "requestedCrit", "requestedExp",
           "ordered", "orderedCrit", "orderedExp",
           "acknowledged", "acknowledgedCrit", "acknowledgedExp":
               #ret := FALSE;
           "idle":
               #ret := TRUE;
       END_CASE;
   END_IF;
   #"Part Request: Validate Remove: Single" := #ret;
END_FUNCTION

FUNCTION "Part Request: Clear Data Table" : Void   // FC48, SCL
{ S7_Optimized_Access := 'TRUE' }
VERSION : 0.1
   VAR_IN_OUT
      dataTable : "Part Request Data";
   END_VAR
   VAR_TEMP
      pRow : Int;
   END_VAR
   VAR CONSTANT
      clearRow : DInt := -1;
   END_VAR
BEGIN
   FOR #pRow := 0 TO "partReqDataRowCount" DO
       #dataTable.row[#pRow] := #clearRow;
   END_FOR;
END_FUNCTION

FUNCTION "Part Request: Collapse Table" : Void   // FC55, SCL
{ S7_Optimized_Access := 'TRUE' }
VERSION : 0.1
   VAR_IN_OUT
      dataTable : "Part Request Data";
   END_VAR
   VAR_TEMP
      pRow : Int;
      pScan : Int;
   END_VAR
BEGIN
   FOR #pRow := 0 TO "partReqDataRowCount" DO
       #pScan := 1;
       IF #dataTable.row[#pRow] <= -1 THEN
           WHILE #dataTable.row[#pRow + #pScan] <= -1 AND #pRow + #pScan < "partReqDataRowCount" DO
               #pScan += 1;
           END_WHILE;
           #dataTable.row[#pRow] := #dataTable.row[#pRow + #pScan];
           #dataTable.row[#pRow + #pScan] := -1;
           IF #pRow + #pScan = "partReqDataRowCount" THEN
               RETURN;
           END_IF;
       END_IF;
   END_FOR;
END_FUNCTION

FUNCTION "Part Request: Validate Remove: WIP" : Bool   // FC89, SCL
{ S7_Optimized_Access := 'TRUE' }
VERSION : 0.1
   VAR_INPUT
      inTable : DInt;
      clearWipRequest : Bool;
   END_VAR
   VAR_TEMP
      ret : Bool;
   END_VAR
BEGIN
   IF #inTable <> -1 THEN
       #ret := #clearWipRequest;
   END_IF;

   #"Part Request: Validate Remove: WIP" := #ret;
END_FUNCTION

// folder: Stations

FUNCTION_BLOCK "Button Parameters"   // FB12, SCL
{ S7_Optimized_Access := 'TRUE' }
VERSION : 0.1
   VAR_INPUT
      pnLib : "Recipe: PN Text Library";
   END_VAR
   VAR_IN_OUT
      stns : "Station: All Stations";
   END_VAR
   VAR
      placeHolder : Bool;
   END_VAR
   VAR_TEMP
      pBtn : Int;
      pStn : Int;
   END_VAR
BEGIN
   REGION "FOR EACH STATION"
       FOR #pStn := 0 TO "STATION_COUNT" DO

           REGION "ON CODE CHANGE"
               IF #stns.stn[#pStn].wipCmpts.flags.newPN THEN

                   REGION "FOR EACH BUTTON"
                       FOR #pBtn := 0 TO "STATION_BUTTON_COUNT" DO

                           REGION "LOAD PARAMETERS"
                               "Load Button Parameters OP"(pnGood := #stns.stn[#pStn].wipCmpts.flags.pnGood[#pBtn],
                                                           btnConfig := #stns.stn[#pStn].kp8Config.btn[#pBtn]);
                           END_REGION

                       END_FOR;
                   END_REGION

               END_IF;
           END_REGION

       END_FOR;
   END_REGION
END_FUNCTION_BLOCK

FUNCTION "Load Button Parameters OP" : Void   // FC2, SCL
{ S7_Optimized_Access := 'TRUE' }
VERSION : 0.1
   VAR_INPUT
      pnGood : Bool;
   END_VAR
   VAR_IN_OUT
      btnConfig : "KP8 Driver: Parameters: 1 Button";
   END_VAR
BEGIN
   REGION "ON GOOD PN"
       IF #pnGood THEN

           REGION "ACTIVATE BUTTON"
               #btnConfig.activate := TRUE;
               #btnConfig.cOff := 'green';
               #btnConfig.cOn1 := 'yellow';
               #btnConfig.cOn2 := '';
               #btnConfig.flash := FALSE;
               #btnConfig.group := 0;
               #btnConfig.mode := TRUE;
           END_REGION

       END_IF;
   END_REGION

   REGION "ON BAD PN"
       IF NOT #pnGood THEN

           REGION "DEACTIVATE BUTTON"
               #btnConfig.activate := FALSE;
               #btnConfig.cOff := 'off';
               #btnConfig.cOn1 := 'off';
               #btnConfig.cOn2 := 'off';
               #btnConfig.flash := FALSE;
               #btnConfig.group := 0;
               #btnConfig.mode := FALSE;
           END_REGION

       END_IF;
   END_REGION
END_FUNCTION

FUNCTION "Expanded Animations" : Void   // FC86, SCL
{ S7_Optimized_Access := 'TRUE' }